VERSION : 0.1
   VAR_INPUT
      OFF_SQ : Bool := false;   // Turn sequence off
      INIT_SQ : Bool := false;   // Set sequence to initial state
      ACK_EF : Bool := false;   // Acknowledge all errors and faults
   END_VAR
   VAR_OUTPUT
      S_NO : Int := 0;   // Step number
      S_MORE : Bool := false;   // More steps are available and can be shown in S_NO
      S_ACTIVE : Bool := false;   // Step indicated in S_NO is active
      ERR_FLT : Bool := false;   // Interlock or supervision group error
      AUTO_ON : Bool := false;   // Automatic mode is active
   END_VAR
   VAR
      HMI_INFO : Array[0..10] of UInt;
      IF_PAR : G7_IfParPlus_V6;
      RT_DATA : G7_RTDataPlus_V6;   // Internal data area
      Abort : G7_TransitionPlus_V6;   // Transition structure
      InitializeTk : G7_TransitionPlus_V6;   // Transition structure
      Block : G7_TransitionPlus_V6;   // Transition structure
      Rdy : G7_TransitionPlus_V6;   // Transition structure
      MixSeq : G7_TransitionPlus_V6;   // Transition structure
      WashSeq : G7_TransitionPlus_V6;   // Transition structure
      Pouring : G7_TransitionPlus_V6;   // Transition structure
      Started : G7_TransitionPlus_V6;   // Transition structure
      Params : G7_TransitionPlus_V6;   // Transition structure
      FillingDn : G7_TransitionPlus_V6;   // Transition structure
      WaterOff : G7_TransitionPlus_V6;   // Transition structure
      TankR : G7_TransitionPlus_V6;   // Transition structure
      "Open Signal_1" : G7_TransitionPlus_V6;   // Transition structure
      MixTimeDn : G7_TransitionPlus_V6;   // Transition structure
      MixOpDn : G7_TransitionPlus_V6;   // Transition structure
      NoFlow : G7_TransitionPlus_V6;   // Transition structure
      MixDn : G7_TransitionPlus_V6;   // Transition structure
      PourSt : G7_TransitionPlus_V6;   // Transition structure
      Rc : G7_TransitionPlus_V6;   // Transition structure
      Transf : G7_TransitionPlus_V6;   // Transition structure
      ClsR : G7_TransitionPlus_V6;   // Transition structure
      Release : G7_TransitionPlus_V6;   // Transition structure
      Init : G7_TransitionPlus_V6;   // Transition structure
      SAut : G7_TransitionPlus_V6;   // Transition structure
      SIn : G7_TransitionPlus_V6;   // Transition structure
      Initd : G7_TransitionPlus_V6;   // Transition structure
      Ab : G7_TransitionPlus_V6;   // Transition structure
      AbortOn : G7_TransitionPlus_V6;   // Transition structure
      DneAbort : G7_TransitionPlus_V6;   // Transition structure
      Idle : G7_StepPlus_V6;   // Step structure
      Ready : G7_StepPlus_V6;   // Step structure
      SelectSeq : G7_StepPlus_V6;   // Step structure
      DoneMix : G7_StepPlus_V6;   // Step structure
      MixStarted : G7_StepPlus_V6;   // Step structure
      "EDIT QWater" : G7_StepPlus_V6;   // Step structure
      FillingUpWater : G7_StepPlus_V6;   // Step structure
      StopReqWater : G7_StepPlus_V6;   // Step structure
      "ReleaseT-104" : G7_StepPlus_V6;   // Step structure
      "USER PourDn" : G7_StepPlus_V6;   // Step structure
      MinMixingTime : G7_StepPlus_V6;   // Step structure
      "USER EndMix" : G7_StepPlus_V6;   // Step structure
      ShuttingDown : G7_StepPlus_V6;   // Step structure
      PouringStarted : G7_StepPlus_V6;   // Step structure
      Recirculation : G7_StepPlus_V6;   // Step structure
      Transfering : G7_StepPlus_V6;   // Step structure
      CloseRoute : G7_StepPlus_V6;   // Step structure
      DoneTransfer : G7_StepPlus_V6;   // Step structure
      StartingInit : G7_StepPlus_V6;   // Step structure
      SetAuto : G7_StepPlus_V6;   // Step structure
      SetInitial : G7_StepPlus_V6;   // Step structure
      Init_Done : G7_StepPlus_V6;   // Step structure
      AbortStarting : G7_StepPlus_V6;   // Step structure
      Aborting : G7_StepPlus_V6;   // Step structure
      Abort_Done : G7_StepPlus_V6;   // Step structure
      SINI : Array[0..3] of USInt;
      LSTT : Array[0..28] of USInt;
      ATAJ : Array[0..28] of USInt;
      ATAB : Array[0..28] of USInt;
      PSTT : Array[0..28] of USInt;
      NSTT : Array[0..28] of USInt;
      ASSJ : Array[0..24] of USInt;
      ASSB : Array[0..24] of USInt;
      PTTS : Array[0..24] of USInt;
      NTTS : Array[0..24] of USInt;
      SW_SQTS : Array[0..24] of USInt;
      SWITCH : Array[0..4] of USInt;
      TVX : Array[0..9] of USInt;
      TTX : Array[0..9] of USInt;
      TSX : Array[0..3] of USInt;
      S00X : Array[0..3] of USInt;
      SOFFX : Array[0..3] of USInt;
      SONX : Array[0..3] of USInt;
      SAX : Array[0..3] of USInt;
      SERRX : Array[0..25] of USInt;
      SMX : Array[0..25] of USInt;
      S0X : Array[0..25] of USInt;
      S1X : Array[0..25] of USInt;
      IL_ALARM_INST : Diag_Alarm;
      SUP_ALARM_INST : Diag_Alarm;
      STEP_TIME_ALARM_INST : Diag_Alarm;
      IEC_TIMER_INST : IEC_TIMER;
      TRANSACTION_FLAG : Bool := false;
   END_VAR
   // LSTT[14] := 255;
   // SINI[0] := 2;
   // SINI[2] := 255;
   // SINI[3] := 255;
   // LSTT[0] := 22;
   // LSTT[1] := 18;
   // LSTT[2] := 255;
   // LSTT[3] := 255;
   // LSTT[4] := 255;
   // LSTT[12] := 255;
   // LSTT[6] := 255;
   // LSTT[7] := 255;
   // LSTT[8] := 255;
   // LSTT[9] := 255;
   // LSTT[10] := 255;
   // LSTT[11] := 255;
   // LSTT[13] := 255;
   // LSTT[15] := 255;
   // LSTT[20] := 255;
   // LSTT[17] := 255;
   // LSTT[18] := 255;
   // LSTT[19] := 255;
   // LSTT[27] := 255;
   // LSTT[22] := 255;
   // LSTT[23] := 255;
   // LSTT[24] := 255;
   // LSTT[25] := 1;
   // LSTT[26] := 255;
   // NSTT[14] := 12;
   // ATAJ[1] := 1;
   // ATAJ[2] := 2;
   // ATAJ[3] := 3;
   // ATAJ[4] := 4;
   // ATAJ[5] := 5;
   // ATAJ[6] := 6;
   // ATAJ[7] := 7;
   // ATAJ[8] := 8;
   // ATAJ[9] := 9;
   // ATAJ[10] := 10;
   // ATAJ[11] := 11;
   // ATAJ[12] := 12;
   // ATAJ[13] := 13;
   // ATAJ[14] := 14;
   // ATAJ[15] := 15;
   // ATAJ[16] := 16;
   // ATAJ[17] := 17;
   // ATAJ[18] := 18;
   // ATAJ[19] := 19;
   // ATAJ[20] := 20;
   // ATAJ[21] := 21;
   // ATAJ[22] := 22;
   // ATAJ[23] := 23;
   // ATAJ[24] := 24;
   // ATAJ[25] := 25;
   // ATAJ[26] := 26;
   // ATAJ[27] := 27;
   // ATAJ[28] := 28;
   // ATAB[0] := 1;
   // ATAB[1] := 2;
   // ATAB[24] := 24;
   // ATAB[3] := 3;
   // ATAB[4] := 5;
   // ATAB[5] := 6;
   // ATAB[6] := 4;
   // ATAB[7] := 7;
   // ATAB[8] := 8;
   // ATAB[9] := 9;
   // ATAB[10] := 10;
   // ATAB[11] := 11;
   // ATAB[12] := 12;
   // ATAB[13] := 13;
   // ATAB[14] := 14;
   // ATAB[15] := 15;
   // ATAB[16] := 16;
   // ATAB[17] := 17;
   // ATAB[18] := 18;
   // ATAB[19] := 19;
   // ATAB[20] := 20;
   // ATAB[21] := 21;
   // ATAB[22] := 22;
   // ATAB[23] := 23;
   // ATAB[25] := 25;
   // ATAB[26] := 26;
   // ATAB[27] := 27;
   // ATAB[28] := 28;
   // PSTT[24] := 20;
   // PSTT[5] := 2;
   // PSTT[3] := 1;
   // PSTT[4] := 2;
   // PSTT[15] := 12;
   // PSTT[6] := 2;
   // PSTT[7] := 4;
   // PSTT[8] := 5;
   // PSTT[9] := 6;
   // PSTT[10] := 7;
   // PSTT[11] := 8;
   // PSTT[12] := 9;
   // PSTT[13] := 10;
   // PSTT[14] := 11;
   // PSTT[16] := 3;
   // PSTT[17] := 13;
   // PSTT[18] := 14;
   // PSTT[19] := 15;
   // PSTT[20] := 16;
   // PSTT[21] := 17;
   // PSTT[22] := 18;
   // PSTT[23] := 19;
   // PSTT[25] := 21;
   // PSTT[26] := 22;
   // PSTT[27] := 23;
   // PSTT[28] := 24;
   // NSTT[0] := 22;
   // NSTT[1] := 18;
   // NSTT[2] := 1;
   // NSTT[3] := 2;
   // NSTT[4] := 4;
   // NSTT[12] := 10;
   // NSTT[6] := 13;
   // NSTT[7] := 5;
   // NSTT[8] := 6;
   // NSTT[9] := 7;
   // NSTT[10] := 8;
   // NSTT[11] := 9;
   // NSTT[13] := 11;
   // NSTT[15] := 3;
   // NSTT[20] := 17;
   // NSTT[17] := 14;
   // NSTT[18] := 15;
   // NSTT[19] := 16;
   // NSTT[27] := 24;
   // NSTT[22] := 19;
   // NSTT[23] := 20;
   // NSTT[24] := 21;
   // NSTT[25] := 1;
   // NSTT[26] := 23;
   // ASSJ[1] := 1;
   // ASSJ[2] := 2;
   // ASSJ[3] := 3;
   // ASSJ[4] := 4;
   // ASSJ[5] := 5;
   // ASSJ[6] := 6;
   // ASSJ[7] := 7;
   // ASSJ[8] := 8;
   // ASSJ[9] := 9;
   // ASSJ[10] := 10;
   // ASSJ[11] := 11;
   // ASSJ[12] := 12;
   // ASSJ[13] := 13;
   // ASSJ[14] := 14;
   // ASSJ[15] := 15;
   // ASSJ[16] := 16;
   // ASSJ[17] := 17;
   // ASSJ[18] := 18;
   // ASSJ[19] := 19;
   // ASSJ[20] := 20;
   // ASSJ[21] := 21;
   // ASSJ[22] := 22;
   // ASSJ[23] := 23;
   // ASSJ[24] := 24;
   // ASSB[1] := 1;
   // ASSB[2] := 2;
   // ASSB[3] := 3;
   // ASSB[4] := 4;
   // ASSB[5] := 5;
   // ASSB[6] := 6;
   // ASSB[7] := 7;
   // ASSB[8] := 8;
   // ASSB[9] := 9;
   // ASSB[10] := 10;
   // ASSB[11] := 11;
   // ASSB[12] := 12;
   // ASSB[13] := 13;
   // ASSB[14] := 14;
   // ASSB[15] := 15;
   // ASSB[16] := 16;
   // ASSB[17] := 17;
   // ASSB[18] := 18;
   // ASSB[19] := 19;
   // ASSB[20] := 20;
   // ASSB[21] := 21;
   // ASSB[22] := 22;
   // ASSB[23] := 23;
   // ASSB[24] := 24;
   // PTTS[0] := 255;
   // PTTS[1] := 2;
   // PTTS[2] := 3;
   // PTTS[3] := 15;
   // PTTS[4] := 4;
   // PTTS[5] := 7;
   // PTTS[6] := 8;
   // PTTS[7] := 9;
   // PTTS[8] := 10;
   // PTTS[9] := 11;
   // PTTS[10] := 12;
   // PTTS[11] := 13;
   // PTTS[12] := 14;
   // PTTS[13] := 6;
   // PTTS[14] := 17;
   // PTTS[15] := 18;
   // PTTS[16] := 19;
   // PTTS[17] := 20;
   // PTTS[18] := 255;
   // PTTS[19] := 22;
   // PTTS[20] := 23;
   // PTTS[21] := 24;
   // PTTS[22] := 255;
   // PTTS[23] := 26;
   // PTTS[24] := 27;
   // NTTS[1] := 3;
   // NTTS[2] := 4;
   // NTTS[3] := 16;
   // NTTS[4] := 7;
   // NTTS[5] := 8;
   // NTTS[6] := 9;
   // NTTS[7] := 10;
   // NTTS[8] := 11;
   // NTTS[9] := 12;
   // NTTS[10] := 13;
   // NTTS[11] := 14;
   // NTTS[12] := 15;
   // NTTS[13] := 17;
   // NTTS[14] := 18;
   // NTTS[15] := 19;
   // NTTS[16] := 20;
   // NTTS[17] := 21;
   // NTTS[18] := 22;
   // NTTS[19] := 23;
   // NTTS[20] := 24;
   // NTTS[21] := 25;
   // NTTS[22] := 26;
   // NTTS[23] := 27;
   // NTTS[24] := 28;
   // SW_SQTS[1] := 1;
   // SW_SQTS[2] := 1;
   // SW_SQTS[3] := 2;
   // SW_SQTS[4] := 2;
   // SW_SQTS[5] := 2;
   // SW_SQTS[6] := 2;
   // SW_SQTS[7] := 2;
   // SW_SQTS[8] := 2;
   // SW_SQTS[9] := 2;
   // SW_SQTS[10] := 2;
   // SW_SQTS[11] := 2;
   // SW_SQTS[12] := 2;
   // SW_SQTS[13] := 3;
   // SW_SQTS[14] := 3;
   // SW_SQTS[15] := 3;
   // SW_SQTS[16] := 3;
   // SW_SQTS[17] := 3;
   // SW_SQTS[18] := 4;
   // SW_SQTS[19] := 4;
   // SW_SQTS[20] := 4;
   // SW_SQTS[21] := 4;
   // SW_SQTS[22] := 5;
   // SW_SQTS[23] := 5;
   // SW_SQTS[24] := 5;
   // SWITCH[0] := 48;
   // SWITCH[1] := 12;
   // SWITCH[2] := 195;
   // SWITCH[3] := 239;
   // SWITCH[4] := 7;
   // TVX[0] := 16#1;
   // TTX[0] := 16#1;
   // TSX[0] := 16#1;
   // S00X[0] := 16#1;
   // SOFFX[0] := 16#1;
   // SONX[0] := 16#1;
   // SAX[0] := 16#1;
   // SERRX[0] := 16#1;
   // SMX[0] := 16#1;
   // S0X[0] := 16#1;
   // S1X[0] := 16#1;
BEGIN
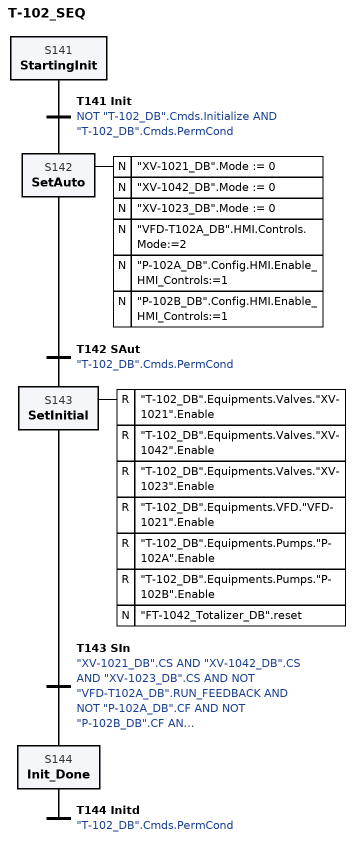
   // permanent pre-instructions
   NETWORK 1
      "T-102_Signals_FROM_R-201"();
      "T-102_Signals_FROM_R-202"();
      "T-102_Signals_FROM_T-104"();
      "T-102_SEQ_FC"();

   // sequencer 1
   STEP StartingInit:   // S141, max time T#10S, warning time T#7S
      // Initialize T-102 Batch sequence
   END_STEP
   TRANSITION Init FROM StartingInit TO SetAuto   // T141
      := NOT "T-102_DB".Cmds.Initialize AND "T-102_DB".Cmds.PermCond;
   END_TRANSITION
   STEP SetAuto:   // S142, max time T#10S, warning time T#7S
              N    "XV-1021_DB".Mode := 0
              N    "XV-1042_DB".Mode := 0
              N    "XV-1023_DB".Mode := 0
              N    "VFD-T102A_DB".HMI.Controls.Mode:=2
              N    "P-102A_DB".Config.HMI.Enable_HMI_Controls:=1
              N    "P-102B_DB".Config.HMI.Enable_HMI_Controls:=1
   END_STEP
   TRANSITION SAut FROM SetAuto TO SetInitial   // T142
      := "T-102_DB".Cmds.PermCond;
   END_TRANSITION
   STEP SetInitial:   // S143, max time T#10S, warning time T#7S
              R    "T-102_DB".Equipments.Valves."XV-1021".Enable
              R    "T-102_DB".Equipments.Valves."XV-1042".Enable
              R    "T-102_DB".Equipments.Valves."XV-1023".Enable
              R    "T-102_DB".Equipments.VFD."VFD-1021".Enable
              R    "T-102_DB".Equipments.Pumps."P-102A".Enable
              R    "T-102_DB".Equipments.Pumps."P-102B".Enable
              N    "FT-1042_Totalizer_DB".reset
   END_STEP
   TRANSITION SIn FROM SetInitial TO Init_Done   // T143
      := "XV-1021_DB".CS AND "XV-1042_DB".CS AND "XV-1023_DB".CS AND NOT "VFD-T102A_DB".RUN_FEEDBACK AND NOT "P-102A_DB".CF AND NOT "P-102B_DB".CF AND ("FT-1042_Totalizer_DB".Total = 0.0) AND "T-102_DB".Cmds.PermCond;
   END_TRANSITION
   STEP Init_Done:   // S144, max time T#10S, warning time T#7S
   END_STEP
   TRANSITION Initd FROM Init_Done TO ?   // T144
      := "T-102_DB".Cmds.PermCond;
   END_TRANSITION

   // permanent post-instructions
   NETWORK 1
      "T-102_FC_Outputs"();
END_FUNCTION_BLOCK

FUNCTION "T-102_SEQ_FC" : Void   // FC76, LAD
{ S7_Optimized_Access := 'TRUE' }
VERSION : 0.1
   VAR_TEMP   // added for the SCL form of the ladder/FBD networks
      _w1 : Bool;
      _w2 : Bool;
      _w3 : Bool;
   END_VAR
BEGIN

REGION Network 2: Abort
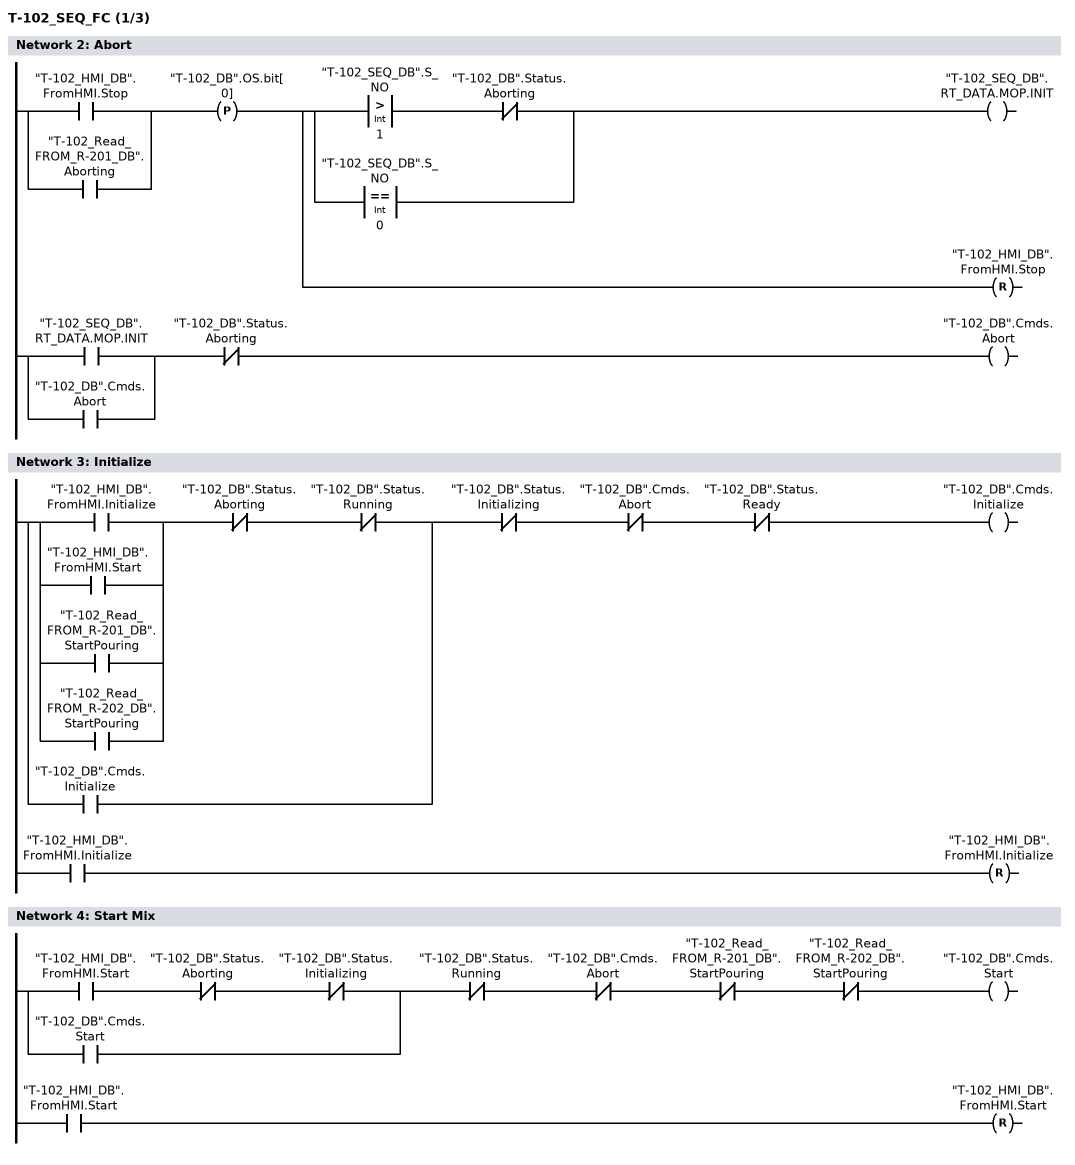
   RUNG wire#powerrail
      Contact( "T-102_HMI_DB".FromHMI.Stop )
      wire#w1
      P_Trig( "T-102_DB".OS.bit[0] )
      wire#w2
      { S7_Templates := "SrcType := Int" } GT_Contact(in1 := "T-102_SEQ_DB".S_NO, in2 := 1)
      I_Contact( "T-102_DB".Status.Aborting )
      wire#w3
      Coil( "T-102_SEQ_DB".RT_DATA.MOP.INIT )
   END_RUNG
   RUNG wire#powerrail
      Contact( "T-102_Read_FROM_R-201_DB".Aborting )
   END_RUNG wire#w1
   RUNG wire#w2
      { S7_Templates := "SrcType := Int" } EQ_Contact(in1 := "T-102_SEQ_DB".S_NO, in2 := 0)
   END_RUNG wire#w3
   RUNG wire#w2
      R_Coil( "T-102_HMI_DB".FromHMI.Stop )
   END_RUNG
   RUNG wire#powerrail
      Contact( "T-102_SEQ_DB".RT_DATA.MOP.INIT )
      wire#w4
      I_Contact( "T-102_DB".Status.Aborting )
      Coil( "T-102_DB".Cmds.Abort )
   END_RUNG
   RUNG wire#powerrail
      Contact( "T-102_DB".Cmds.Abort )
   END_RUNG wire#w4
   // the same network as SCL:
   #_w1 := "T-102_HMI_DB".FromHMI.Stop OR "T-102_Read_FROM_R-201_DB".Aborting;
   #_w2 := #_w1 AND NOT "T-102_DB".OS.bit[0];   // rising edge
   "T-102_DB".OS.bit[0] := #_w1;
   "T-102_SEQ_DB".RT_DATA.MOP.INIT := #_w2 AND ((("T-102_SEQ_DB".S_NO > 1) AND NOT "T-102_DB".Status.Aborting) OR ("T-102_SEQ_DB".S_NO = 0));
   IF #_w2 THEN "T-102_HMI_DB".FromHMI.Stop := FALSE; END_IF;
   "T-102_DB".Cmds.Abort := ("T-102_SEQ_DB".RT_DATA.MOP.INIT OR "T-102_DB".Cmds.Abort) AND NOT "T-102_DB".Status.Aborting;
END_REGION

REGION Network 3: Initialize
   RUNG wire#powerrail
      Contact( "T-102_HMI_DB".FromHMI.Initialize )
      wire#w1
      I_Contact( "T-102_DB".Status.Aborting )
      I_Contact( "T-102_DB".Status.Running )
      wire#w2
      I_Contact( "T-102_DB".Status.Initializing )
      I_Contact( "T-102_DB".Cmds.Abort )
      I_Contact( "T-102_DB".Status.Ready )
      Coil( "T-102_DB".Cmds.Initialize )
   END_RUNG
   RUNG wire#powerrail
      Contact( "T-102_HMI_DB".FromHMI.Start )
   END_RUNG wire#w1
   RUNG wire#powerrail
      Contact( "T-102_Read_FROM_R-201_DB".StartPouring )
   END_RUNG wire#w1
   RUNG wire#powerrail
      Contact( "T-102_Read_FROM_R-202_DB".StartPouring )
   END_RUNG wire#w1
   RUNG wire#powerrail
      Contact( "T-102_DB".Cmds.Initialize )
   END_RUNG wire#w2
   RUNG wire#powerrail
      Contact( "T-102_HMI_DB".FromHMI.Initialize )
      R_Coil( "T-102_HMI_DB".FromHMI.Initialize )
   END_RUNG
   // the same network as SCL:
   "T-102_DB".Cmds.Initialize := ((("T-102_HMI_DB".FromHMI.Initialize OR "T-102_HMI_DB".FromHMI.Start OR "T-102_Read_FROM_R-201_DB".StartPouring OR "T-102_Read_FROM_R-202_DB".StartPouring) AND NOT "T-102_DB".Status.Aborting AND NOT "T-102_DB".Status.Running) OR "T-102_DB".Cmds.Initialize) AND NOT "T-102_DB".Status.Initializing AND NOT "T-102_DB".Cmds.Abort AND NOT "T-102_DB".Status.Ready;
   IF "T-102_HMI_DB".FromHMI.Initialize THEN "T-102_HMI_DB".FromHMI.Initialize := FALSE; END_IF;
END_REGION

REGION Network 4: Start Mix
   RUNG wire#powerrail
      Contact( "T-102_HMI_DB".FromHMI.Start )
      I_Contact( "T-102_DB".Status.Aborting )
      I_Contact( "T-102_DB".Status.Initializing )
      wire#w1
      I_Contact( "T-102_DB".Status.Running )
      I_Contact( "T-102_DB".Cmds.Abort )
      I_Contact( "T-102_Read_FROM_R-201_DB".StartPouring )
      I_Contact( "T-102_Read_FROM_R-202_DB".StartPouring )
      Coil( "T-102_DB".Cmds.Start )
   END_RUNG
   RUNG wire#powerrail
      Contact( "T-102_DB".Cmds.Start )
   END_RUNG wire#w1
   RUNG wire#powerrail
      Contact( "T-102_HMI_DB".FromHMI.Start )
      R_Coil( "T-102_HMI_DB".FromHMI.Start )
   END_RUNG
   // the same network as SCL:
   "T-102_DB".Cmds.Start := (("T-102_HMI_DB".FromHMI.Start AND NOT "T-102_DB".Status.Aborting AND NOT "T-102_DB".Status.Initializing) OR "T-102_DB".Cmds.Start) AND NOT "T-102_DB".Status.Running AND NOT "T-102_DB".Cmds.Abort AND NOT "T-102_Read_FROM_R-201_DB".StartPouring AND NOT "T-102_Read_FROM_R-202_DB".StartPouring;
   IF "T-102_HMI_DB".FromHMI.Start THEN "T-102_HMI_DB".FromHMI.Start := FALSE; END_IF;
END_REGION

REGION Network 5: Procedure Selected
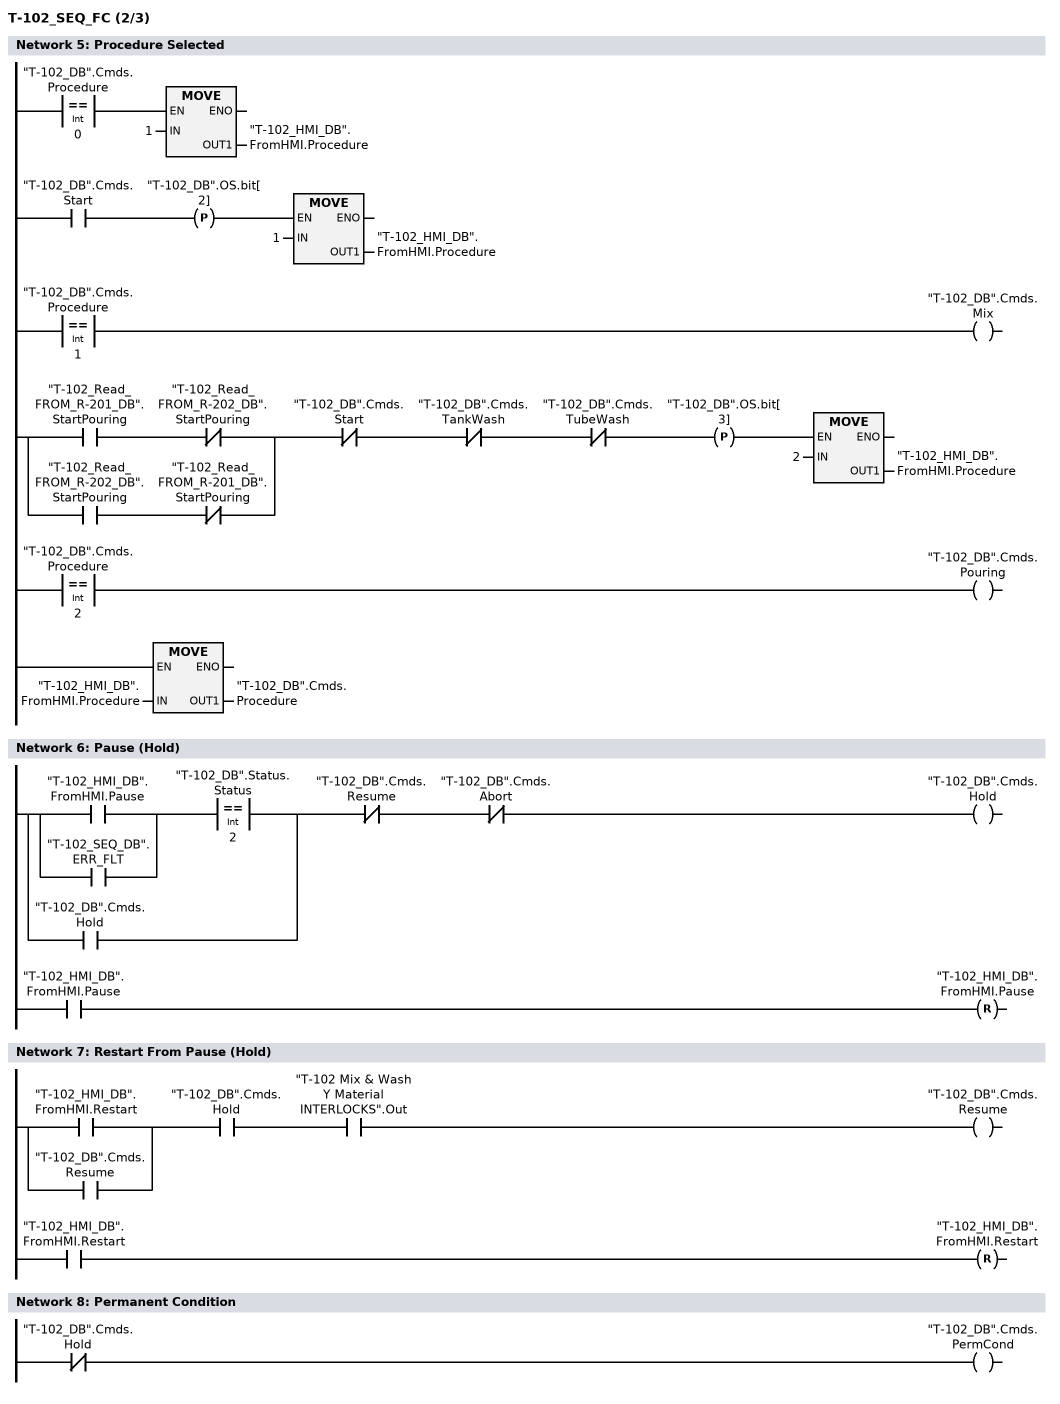
   RUNG wire#powerrail
      { S7_Templates := "SrcType := Int" } EQ_Contact(in1 := "T-102_DB".Cmds.Procedure, in2 := 0)
      Move(in := 1, out1 => "T-102_HMI_DB".FromHMI.Procedure)
   END_RUNG
   RUNG wire#powerrail
      Contact( "T-102_DB".Cmds.Start )
      P_Trig( "T-102_DB".OS.bit[2] )
      Move(in := 1, out1 => "T-102_HMI_DB".FromHMI.Procedure)
   END_RUNG
   RUNG wire#powerrail
      { S7_Templates := "SrcType := Int" } EQ_Contact(in1 := "T-102_DB".Cmds.Procedure, in2 := 1)
      Coil( "T-102_DB".Cmds.Mix )
   END_RUNG
   RUNG wire#powerrail
      Contact( "T-102_Read_FROM_R-201_DB".StartPouring )
      I_Contact( "T-102_Read_FROM_R-202_DB".StartPouring )
      wire#w1
      I_Contact( "T-102_DB".Cmds.Start )
      I_Contact( "T-102_DB".Cmds.TankWash )
      I_Contact( "T-102_DB".Cmds.TubeWash )
      P_Trig( "T-102_DB".OS.bit[3] )
      Move(in := 2, out1 => "T-102_HMI_DB".FromHMI.Procedure)
   END_RUNG
   RUNG wire#powerrail
      Contact( "T-102_Read_FROM_R-202_DB".StartPouring )
      I_Contact( "T-102_Read_FROM_R-201_DB".StartPouring )
   END_RUNG wire#w1
   RUNG wire#powerrail
      { S7_Templates := "SrcType := Int" } EQ_Contact(in1 := "T-102_DB".Cmds.Procedure, in2 := 2)
      Coil( "T-102_DB".Cmds.Pouring )
   END_RUNG
   RUNG wire#powerrail
      Move(in := "T-102_HMI_DB".FromHMI.Procedure, out1 => "T-102_DB".Cmds.Procedure)
   END_RUNG
   // the same network as SCL:
   IF "T-102_DB".Cmds.Procedure = 0 THEN "T-102_HMI_DB".FromHMI.Procedure := 1; END_IF;
   #_w1 := "T-102_DB".Cmds.Start AND NOT "T-102_DB".OS.bit[2];   // rising edge
   "T-102_DB".OS.bit[2] := "T-102_DB".Cmds.Start;
   IF #_w1 THEN "T-102_HMI_DB".FromHMI.Procedure := 1; END_IF;
   "T-102_DB".Cmds.Mix := "T-102_DB".Cmds.Procedure = 1;
   #_w2 := (("T-102_Read_FROM_R-201_DB".StartPouring AND NOT "T-102_Read_FROM_R-202_DB".StartPouring) OR ("T-102_Read_FROM_R-202_DB".StartPouring AND NOT "T-102_Read_FROM_R-201_DB".StartPouring)) AND NOT "T-102_DB".Cmds.Start AND NOT "T-102_DB".Cmds.TankWash AND NOT "T-102_DB".Cmds.TubeWash;
   #_w3 := #_w2 AND NOT "T-102_DB".OS.bit[3];   // rising edge
   "T-102_DB".OS.bit[3] := #_w2;
   IF #_w3 THEN "T-102_HMI_DB".FromHMI.Procedure := 2; END_IF;
   "T-102_DB".Cmds.Pouring := "T-102_DB".Cmds.Procedure = 2;
   "T-102_DB".Cmds.Procedure := "T-102_HMI_DB".FromHMI.Procedure;
END_REGION

REGION Network 6: Pause (Hold)
   RUNG wire#powerrail
      Contact( "T-102_HMI_DB".FromHMI.Pause )
      wire#w1
      { S7_Templates := "SrcType := Int" } EQ_Contact(in1 := "T-102_DB".Status.Status, in2 := 2)
      wire#w2
      I_Contact( "T-102_DB".Cmds.Resume )
      I_Contact( "T-102_DB".Cmds.Abort )
      Coil( "T-102_DB".Cmds.Hold )
   END_RUNG
   RUNG wire#powerrail
      Contact( "T-102_SEQ_DB".ERR_FLT )
   END_RUNG wire#w1
   RUNG wire#powerrail
      Contact( "T-102_DB".Cmds.Hold )
   END_RUNG wire#w2
   RUNG wire#powerrail
      Contact( "T-102_HMI_DB".FromHMI.Pause )
      R_Coil( "T-102_HMI_DB".FromHMI.Pause )
   END_RUNG
   // the same network as SCL:
   "T-102_DB".Cmds.Hold := ((("T-102_HMI_DB".FromHMI.Pause OR "T-102_SEQ_DB".ERR_FLT) AND ("T-102_DB".Status.Status = 2)) OR "T-102_DB".Cmds.Hold) AND NOT "T-102_DB".Cmds.Resume AND NOT "T-102_DB".Cmds.Abort;
   IF "T-102_HMI_DB".FromHMI.Pause THEN "T-102_HMI_DB".FromHMI.Pause := FALSE; END_IF;
END_REGION

REGION Network 7: Restart From Pause (Hold)
   RUNG wire#powerrail
      Contact( "T-102_HMI_DB".FromHMI.Restart )
      wire#w1
      Contact( "T-102_DB".Cmds.Hold )
      Contact( "T-102 Mix & Wash Y Material  INTERLOCKS".Out )
      Coil( "T-102_DB".Cmds.Resume )
   END_RUNG
   RUNG wire#powerrail
      Contact( "T-102_DB".Cmds.Resume )
   END_RUNG wire#w1
   RUNG wire#powerrail
      Contact( "T-102_HMI_DB".FromHMI.Restart )
      R_Coil( "T-102_HMI_DB".FromHMI.Restart )
   END_RUNG
   // the same network as SCL:
   "T-102_DB".Cmds.Resume := ("T-102_HMI_DB".FromHMI.Restart OR "T-102_DB".Cmds.Resume) AND "T-102_DB".Cmds.Hold AND "T-102 Mix & Wash Y Material  INTERLOCKS".Out;
   IF "T-102_HMI_DB".FromHMI.Restart THEN "T-102_HMI_DB".FromHMI.Restart := FALSE; END_IF;
END_REGION

REGION Network 8: Permanent Condition
   RUNG wire#powerrail
      I_Contact( "T-102_DB".Cmds.Hold )
      Coil( "T-102_DB".Cmds.PermCond )
   END_RUNG
   // the same network as SCL:
   "T-102_DB".Cmds.PermCond := NOT "T-102_DB".Cmds.Hold;
END_REGION

REGION Network 9: Tank Wash
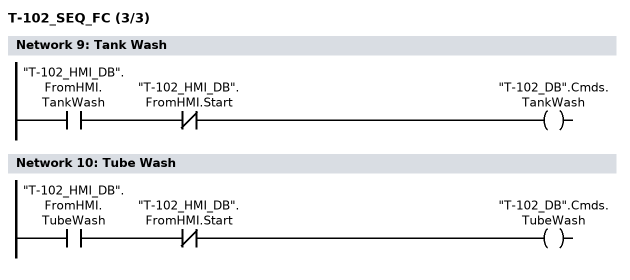
   RUNG wire#powerrail
      Contact( "T-102_HMI_DB".FromHMI.TankWash )
      I_Contact( "T-102_HMI_DB".FromHMI.Start )
      Coil( "T-102_DB".Cmds.TankWash )
   END_RUNG
   // the same network as SCL:
   "T-102_DB".Cmds.TankWash := "T-102_HMI_DB".FromHMI.TankWash AND NOT "T-102_HMI_DB".FromHMI.Start;
END_REGION

REGION Network 10: Tube Wash
   RUNG wire#powerrail
      Contact( "T-102_HMI_DB".FromHMI.TubeWash )
      I_Contact( "T-102_HMI_DB".FromHMI.Start )
      Coil( "T-102_DB".Cmds.TubeWash )
   END_RUNG
   // the same network as SCL:
   "T-102_DB".Cmds.TubeWash := "T-102_HMI_DB".FromHMI.TubeWash AND NOT "T-102_HMI_DB".FromHMI.Start;
END_REGION

REGION Network 11 (SCL): Sequence Status
   IF "T-102_SEQ_DB".S_NO= 1 THEN
       "T-102_DB".Status.Status := 1; //Idle
   ELSIF "T-102_SEQ_DB".S_NO > 1 AND "T-102_SEQ_DB".S_NO < 150  AND NOT "T-102_SEQ_DB".ERR_FLT AND NOT "T-102_DB".Cmds.Hold THEN
       "T-102_DB".Status.Status := 2; //Running
   ELSIF "T-102_SEQ_DB".S_NO >= 151 AND "T-102_SEQ_DB".S_NO <= 160 AND NOT "T-102_SEQ_DB".ERR_FLT THEN
       "T-102_DB".Status.Status := 3; // Stopping
   ELSIF "T-102_SEQ_DB".ERR_FLT  AND  ("T-102_SEQ_DB".S_NO > 1 AND "T-102_SEQ_DB".S_NO < 150) THEN
       "T-102_DB".Status.Status := 4; //Held
   ELSIF  "T-102_SEQ_DB".ERR_FLT AND  ("T-102_SEQ_DB".S_NO > 1 AND "T-102_SEQ_DB".S_NO < 150) AND "T-102_Aux_DB"."Bool".TOff  THEN
       "T-102_DB".Status.Status := 5; // Holding
   ELSE
       "T-102_DB".Status.Status := 6; //Unknown
   END_IF;

   "T-102_DB".Status.Running := ("T-102_SEQ_DB".S_NO > 3 AND "T-102_SEQ_DB".S_NO <= 150);
   "T-102_DB".Status.Initializing := ("T-102_SEQ_DB".S_NO >= 141 AND "T-102_SEQ_DB".S_NO <= 150);

   //Enable/Disable HMI Start/Stop Button
   "T-102_HMI_DB".ToHMI.EnStopButton := ("T-102_DB".Status.Status > 1) OR "T-102_DB".Status.Step = 0; //Enable HMI Stop Button
   "T-102_HMI_DB".ToHMI.EnStartButton := "T-102_DB".Status.Status = 1; //Enable Start Button
   "T-102_HMI_DB".ToHMI.EnPauseButton := "T-102_DB".Status.Status = 2; //Enable Pause Button
   "T-102_HMI_DB".ToHMI.EnRestartButton := "T-102_DB".Status.Status = 4; //Enable Pause Button

   //****Interlock Activated
   "T-102_HMI_DB".ToHMI.InterlockActivated := "T-102 Mix & Wash Y Material  INTERLOCKS".Out;
END_REGION

REGION Network 12 (SCL): Sequence Step
   "T-102_DB".Status.Step := "T-102_SEQ_DB".S_NO;
END_REGION

REGION Network 13 (SCL): Sequence state (Procedure running)
   IF "T-102_SEQ_DB".S_NO = 3 OR "T-102_SEQ_DB".S_NO = 4 THEN
       "T-102_DB".Status.State := 1; //Ready
   ELSIF "T-102_SEQ_DB".S_NO >= 21 AND "T-102_SEQ_DB".S_NO <= 60 THEN
       "T-102_DB".Status.State := 2; //Mixing 
   ELSIF "T-102_SEQ_DB".S_NO >= 61 AND "T-102_SEQ_DB".S_NO <= 80 THEN
       "T-102_DB".Status.State := 3; //Pouring
   ELSIF "T-102_SEQ_DB".S_NO >= 141 AND "T-102_SEQ_DB".S_NO <= 150 THEN
       "T-102_DB".Status.State := 4; //Initializing
   ELSIF "T-102_SEQ_DB".S_NO >= 151 AND "T-102_SEQ_DB".S_NO <= 160 THEN
       "T-102_DB".Status.State := 5; //Aborting
   ELSE
       "T-102_DB".Status.State := 0;
   END_IF;
END_REGION

REGION Network 14: Sequence State
END_REGION
END_FUNCTION

FUNCTION "T-102_FC_Outputs" : Void   // FC83, SCL
{ S7_Optimized_Access := 'TRUE' }
VERSION : 0.1
   VAR_TEMP
      Pump_A : Struct
         Cond_01 : Bool;   // Condition 01
         Cond_02 : Bool;
         Cond_03 : Bool;   // Condition 03
      END_STRUCT;
      Pump_B : Struct
         Cond_01 : Bool;   // Condition 01
         Cond_02 : Bool;   // Condition 02
         Cond_03 : Bool;   // Condition 03
      END_STRUCT;
      XV : Struct
         "1021" : Bool;
         "1042" : Bool;
         "1023" : Bool;
      END_STRUCT;
      RouteOpened : Bool;
      PumpsOff : Bool;
      Recirculating : Bool;
   END_VAR
BEGIN
   //****** Equipmens Activation*******
   //
   //**************************************************************
   //
   //
   //IF "AlwaysFALSE" THEN
       //***********************************************Tank Outlet Valve**********************************************************************
       IF "XV-1021_DB".Mode = 0 THEN
           "T-102_DB".Equipments.Valves."XV-1021".CmdOn := "T-102_DB".Equipments.Valves."XV-1021".Enable AND NOT "T-102_DB".Cmds.Hold;
           //Delay Off To avoid Overpressure the Lines
           #XV."1021" := "T-102_DB".Equipments.Valves."XV-1021".CmdOn;
           "T-102_Aux_DB".Timer."XV-1021".TOF(IN := #XV."1021",
                                              PT := "T-102_Aux_DB".Constants.CmdDelay);
           //Command to the Valve
           IF "T-102_Aux_DB".Timer."XV-1021".Q THEN
               "XV-1021_DB".CMD := 2;
           ELSE
               "XV-1021_DB".CMD := 1;
           END_IF;
           "T-102_DB".Equipments.Valves."XV-1021".TurningOff := NOT "T-102_DB".Equipments.Valves."XV-1021".CmdOn AND "T-102_Aux_DB".Timer."XV-1021".Q;
       END_IF;
       //***********************************************Tank Inlet Valve**********************************************************************
       IF "XV-1042_DB".Mode = 0 THEN
           "T-102_DB".Equipments.Valves."XV-1042".CmdOn := "T-102_DB".Equipments.Valves."XV-1042".Enable AND NOT "T-102_DB".Cmds.Hold;
           //Delay Off To avoid Overpressure the Lines
           #XV."1042" := "T-102_DB".Equipments.Valves."XV-1042".CmdOn;
           "T-102_Aux_DB".Timer."XV-1042".TOF(IN := #XV."1042",
                                              PT := "T-102_Aux_DB".Constants.CmdDelay);
           //Command to the Valve
           IF "T-102_Aux_DB".Timer."XV-1042".Q THEN
               "XV-1042_DB".CMD := 2;
           ELSE
               "XV-1042_DB".CMD := 1;
           END_IF;
           "T-102_DB".Equipments.Valves."XV-1042".TurningOff := NOT "T-102_DB".Equipments.Valves."XV-1042".CmdOn AND "T-102_Aux_DB".Timer."XV-1042".Q;
       END_IF;
       //***********************************************Tank Transfer Valve**********************************************************************
       IF "XV-1023_DB".Mode = 0 THEN
           "T-102_DB".Equipments.Valves."XV-1023".CmdOn := "T-102_DB".Equipments.Valves."XV-1023".Enable AND NOT "T-102_DB".Cmds.Hold;
           //Delay Off To avoid Overpressure the Lines
           #XV."1023" := "T-102_DB".Equipments.Valves."XV-1023".CmdOn;
           "T-102_Aux_DB".Timer."XV-1023".TOF(IN := #XV."1023",
                                              PT := "T-102_Aux_DB".Constants.CmdDelay);
           //Command to the Valve
           IF "T-102_Aux_DB".Timer."XV-1023".Q THEN
               "XV-1023_DB".CMD := 2;
           ELSE
               "XV-1023_DB".CMD := 1;
           END_IF;
           "T-102_DB".Equipments.Valves."XV-1023".TurningOff := NOT "T-102_DB".Equipments.Valves."XV-1023".CmdOn AND "T-102_Aux_DB".Timer."XV-1023".Q;
       END_IF;
       //***********************************************Feed Water Pump A**********************************************************************
       // Condition to CmdOn "On Command" 
       IF "P-102A_DB".Config.HMI.Enable_HMI_Controls = 1 THEN
           #Pump_A.Cond_01 := "T-102_DB".Equipments.Pumps."P-102A".Enable AND ("T-102_DB".PmpSel."P-102AB" = 1 OR "T-102_DB".PmpSel."P-102AB" = 3);
           #Pump_A.Cond_02 := "T-102_Write_TO_R-201_DB".RouteOpened AND "T-102_Read_FROM_R-201_DB".RouteOpened OR ("T-102_Write_TO_R-202_DB".RouteOpened AND "T-102_Read_FROM_R-202_DB".RouteOpened); //Route Open to sent to the Reactor
           #Pump_A.Cond_03 := "XV-1021_DB".OS AND "XV-1023_DB".CS; //Route open to Recirculate
           "T-102_DB".Equipments.Pumps."P-102A".CmdOn := #Pump_A.Cond_01 AND (#Pump_A.Cond_02 OR #Pump_A.Cond_03) AND NOT "T-102_DB".Cmds.Hold;
           IF "T-102_DB".Equipments.Pumps."P-102A".CmdOn THEN
               "P-102A_DB".Stop_CMD := False;
               "P-102A_DB".Start_CMD := true;
               "P-102A_DB".ON := TRUE;
               "P-102A_DB".OFF := FALSE;
           ELSE
               "P-102A_DB".Stop_CMD := True;
               "P-102A_DB".Start_CMD := False;
               "P-102A_DB".ON := FALSE;
               "P-102A_DB".OFF := TRUE;
           END_IF;
       END_IF;

       //***********************************************Feed Water Pump B**********************************************************************
       // Condition to CmdOn "On Command" 
       IF "P-102B_DB".Config.HMI.Enable_HMI_Controls = 1 THEN
           #Pump_B.Cond_01 := "T-102_DB".Equipments.Pumps."P-102B".Enable AND ("T-102_DB".PmpSel."P-102AB" = 2 OR "T-102_DB".PmpSel."P-102AB" = 3);
           #Pump_B.Cond_02 := "T-102_Write_TO_R-201_DB".RouteOpened AND "T-102_Read_FROM_R-201_DB".RouteOpened  OR ("T-102_Write_TO_R-202_DB".RouteOpened AND "T-102_Read_FROM_R-202_DB".RouteOpened); //Route Open to sent to the Reactor
           #Pump_B.Cond_03 := "XV-1021_DB".OS AND "XV-1023_DB".CS; //Route open to Recirculate
           "T-102_DB".Equipments.Pumps."P-102B".CmdOn := #Pump_B.Cond_01 AND (#Pump_B.Cond_02 OR #Pump_B.Cond_03) AND NOT "T-102_DB".Cmds.Hold;
           IF "T-102_DB".Equipments.Pumps."P-102B".CmdOn THEN
               "P-102B_DB".Stop_CMD := False;
               "P-102B_DB".Start_CMD := true;
               "P-102B_DB".ON := TRUE;
               "P-102B_DB".OFF := FALSE;
           ELSE
               "P-102B_DB".Stop_CMD := True;
               "P-102B_DB".Start_CMD := False;
               "P-102B_DB".ON := FALSE;
               "P-102B_DB".OFF := TRUE;
           END_IF;
       END_IF;
       //***********************************************Mixer***********************************************************************
       IF "VFD-T102A_DB".HMI.Controls.Mode = 2 THEN
           "T-102_DB".Equipments.VFD."VFD-1021".CmdOn := "T-102_DB".Equipments.VFD."VFD-1021".Enable AND NOT "T-102_DB".Cmds.Hold;
           IF "T-102_DB".Equipments.VFD."VFD-1021".CmdOn THEN
               "VFD-T102A_DB".PLCCommand := TRUE;
           ELSE
               "VFD-T102A_DB".PLCCommand := FALSE;
           END_IF;
       END_IF;
   //END_IF;

   //Interlocks Signals to R-201
   //*****Recirculating*****//
   #Recirculating := ("P-102A_DB".CF OR "P-102B_DB".CF) AND ("XV-1021_DB".OS AND "XV-1023_DB".CS) AND ("FT-1021_DB".SAI > 0.2);

   "T-102_Write_TO_R-201_DB".Recirculating :=   #Recirculating;
   "T-102_Write_TO_R-202_DB".Recirculating :=   #Recirculating;
   //****Route open to Reactors*****//
   #RouteOpened := "XV-1021_DB".OS AND "XV-1023_DB".OS;

   "T-102_Write_TO_R-201_DB".RouteOpened :=  #RouteOpened ;
   "T-102_Write_TO_R-202_DB".RouteOpened :=  #RouteOpened ;
   //*****Pumps OFF*****//
   #PumpsOff := NOT "P-102A_DB".CF AND NOT "P-102B_DB".CF AND ("PT-102A_DB".SAI < 0.8 AND "PT-102B_DB".SAI < 0.8);

   "T-102_Write_TO_R-201_DB".PupmsOFF :=#PumpsOff ;
   "T-102_Write_TO_R-202_DB".PupmsOFF := #PumpsOff ;

       //********************Pouring Status*********************************
   "T-102_DB".Status.PouringRunning := ("T-102_DB".Status.Step = 61 OR "T-102_DB".Status.Step = 62 OR "T-102_DB".Status.Step = 63) AND (#RouteOpened AND NOT #PumpsOff);

   //***************Interlocks to T-104***************//
   "T-102_Write_TO_T-104_DB".ReqWaterToMix := "XV-1042_DB".OS AND "T-102_DB".ExchangeCmds.Send.ReqWater;
   "T-102_Write_TO_T-104_DB".StopReqWaterToMix := "T-102_DB".ExchangeCmds.Send.StopReqWater;

   //***************Valves Status***************//
   "T-102_Aux_DB"."Bool".TOff := "T-102_DB".Equipments.Valves."XV-1021".TurningOff OR "T-102_DB".Equipments.Valves."XV-1042".TurningOff OR "T-102_DB".Equipments.Valves."XV-1023".TurningOff;
   //***************Timer***************//
   "T-102_Aux_DB"."Bool".MinMixT_Enab := "T-102_DB".Status.Step = 27 AND "VFD-T102A_DB".RUN_FEEDBACK AND "VFD-T102A_DB".SPEED_FEEDBACK > 500;
   "T-102_Aux_DB"."Bool".MinMixT_Reset := "T-102_DB".Cmds.Abort OR "T-102_DB".Status.Step = 1;
END_FUNCTION

// folder: State MACHINE/1)Tanks/Tank T-102 (Y)/T-102 <---> R-201

FUNCTION "T-102_Signals_FROM_R-201" : Void   // FC64, LAD
{ S7_Optimized_Access := 'TRUE' }
VERSION : 0.1
BEGIN

REGION Network 1: Start Pouring Sequence
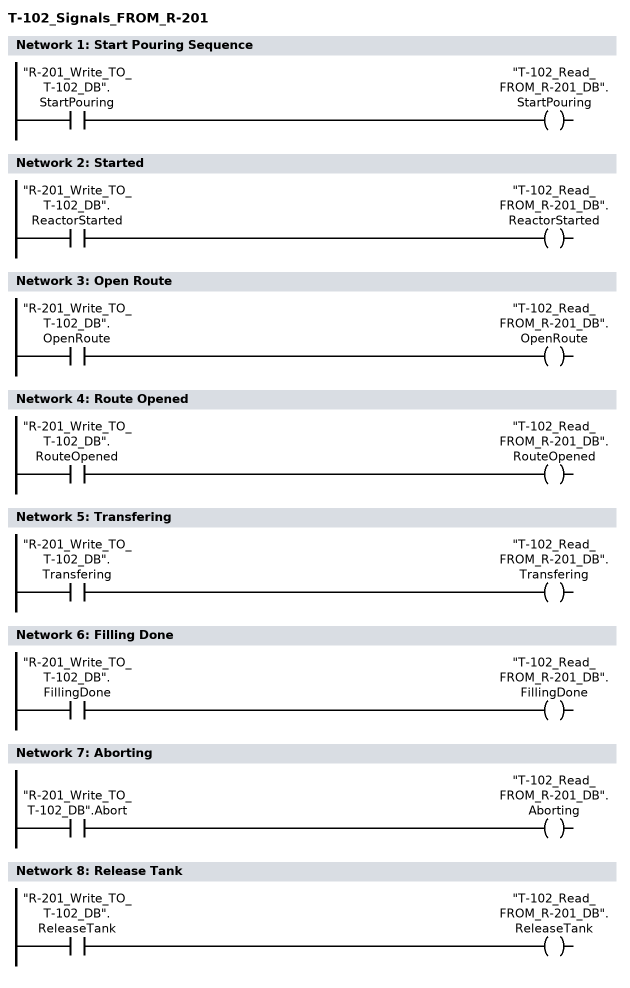
   RUNG wire#powerrail
      Contact( "R-201_Write_TO_T-102_DB".StartPouring )
      Coil( "T-102_Read_FROM_R-201_DB".StartPouring )
   END_RUNG
   // the same network as SCL:
   "T-102_Read_FROM_R-201_DB".StartPouring := "R-201_Write_TO_T-102_DB".StartPouring;
END_REGION

REGION Network 2: Started
   RUNG wire#powerrail
      Contact( "R-201_Write_TO_T-102_DB".ReactorStarted )
      Coil( "T-102_Read_FROM_R-201_DB".ReactorStarted )
   END_RUNG
   // the same network as SCL:
   "T-102_Read_FROM_R-201_DB".ReactorStarted := "R-201_Write_TO_T-102_DB".ReactorStarted;
END_REGION

REGION Network 3: Open Route
   RUNG wire#powerrail
      Contact( "R-201_Write_TO_T-102_DB".OpenRoute )
      Coil( "T-102_Read_FROM_R-201_DB".OpenRoute )
   END_RUNG
   // the same network as SCL:
   "T-102_Read_FROM_R-201_DB".OpenRoute := "R-201_Write_TO_T-102_DB".OpenRoute;
END_REGION

REGION Network 4: Route Opened
   RUNG wire#powerrail
      Contact( "R-201_Write_TO_T-102_DB".RouteOpened )
      Coil( "T-102_Read_FROM_R-201_DB".RouteOpened )
   END_RUNG
   // the same network as SCL:
   "T-102_Read_FROM_R-201_DB".RouteOpened := "R-201_Write_TO_T-102_DB".RouteOpened;
END_REGION
